
     #BLEND:
       // ========================================================================================================
       // Blending 
       // ========================================================================================================
       // Definition of blending (PathData: cmdParameters.bufferMode)
       // The parameter name is defined as "BLEND"
       // 
       // If "BLEND" was found, set the defined values in the connected PathData
       // The values are defined as "DirectValues" because the value to set is directly written here in this FC
       // Buffer mode (cmdParameters.bufferMode)
       // #parameterDefinition.directValues.cmdParameters.bufferMode := 5;
       // --> Set the bufferMode to 5 (Blending with high velocity)
       // 
       // Also set the priority #parameterDefinition.priorities.cmdParameters.bufferMode := "LKINLANG_PRIO_DEFINED";
       // 
       // Properties:
       // ----------
       // "LKINLANG_PRG_MODAL": Modal in program to save velocity value once set
       // 
       // Conditions:
       // ----------
       // Conditions are used to make other parameters mandatory.
       // Here the parameter "RADIUS" must be programmed the same line, because blending consits of the bufferMode and the TransitionParameter[1].
       // There can be up to "LKINLANG_NUMBER_OF_CONDITIONS" conditions.
       // How to configure:
       // 1. Set conditions[#tempConditionCounter].ParameterNumber to the parameter you want to check
       // 2. Set conditions[#tempConditionCounter].Mode according to where the parameter has to be written
       //    These modes are possible:
       //    "LKINLANG_CONDITION_IN_LINE" --> Selected parameter must be written in the same line
       //    "LKINLANG_CONDITION_IN_COMMAND" --> Selected parameter must be written in the same motion command
       //    "LKINLANG_CONDITION_IN_PROGRAM" --> Selected parameter must be written somewhere in the program before
       // 3. The setting #parameterDefinition.conditions[#tempConditionCounter].Group can be used to group parameters
       //    Only one condition of each group must be fulfilled.
       //    Also make sure groups are not used twice for other parameters; they must be unique
       //    
       // 
       // Parameter name definition
       #parameterDefinition.parameterNameString := 'BLEND';
       #parameterDefinition.parameterNameNumber := -1;

       // Matching to PathData
       #parameterDefinition.directValues.cmdParameters.bufferMode := 5; // BlendHigh

       // Priorities
       #parameterDefinition.priorities.cmdParameters.bufferMode := "LKINLANG_PRIO_DEFINED";

       // Properties
       #parameterDefinition.properties := "LKINLANG_PRG_MODAL";

       // Conditions
       #tempConditionCounter := 1;
       #parameterDefinition.conditions[#tempConditionCounter].ParameterNumber := #RADIUS;
       #parameterDefinition.conditions[#tempConditionCounter].Mode := "LKINLANG_CONDITION_IN_LINE";
       #parameterDefinition.conditions[#tempConditionCounter].Group := 10;

       // Valid counts per line
       #parameterDefinition.validCountPerLine := 1;
       // ========================================================================================================


     #RADIUS:
       // ========================================================================================================
       // Transition parameter
       // ========================================================================================================
       // Definition of TransitionParameter[1] (PathData: cmdParameters.transitionParameters[1])
       // The parameter name is defined as "R"
       // 
       // If "R" was found, set the defined values in the connected PathData
       // The value is defined as "FollowingValue" because the value is not written here, but in the program line after this parameter
       // e.g. R15 <-- 15 is taken as transitionParameter[1]
       // To do this, set #parameterDefinition.followingValues[1].cmdParameters.transitionParameters[1] := TRUE;
       // 
       // Also set the priority #parameterDefinition.priorities.cmdParameters.transitionParameters[1] := "LKINLANG_PRIO_DEFINED";
       // 
       // Properties:
       // ----------
       // "LKINLANG_PRG_MODAL": Modal in program to save transition parameter
       // 
       // Conditions:
       // ----------
       // This parameter is a condition for "BLEND", whenever "BLEND" is programmed, also "R" must be written in the same line.
       // See definition above.
       // 
       //
       // Parameter name definition
       #parameterDefinition.parameterNameString := 'R';
       #parameterDefinition.parameterNameNumber := -1;

       // Matching to PathData
       #parameterDefinition.followingValues[1].cmdParameters.transitionParameters[1] := TRUE; // Transition parameter [1] is set

       // Priorities
       #parameterDefinition.priorities.cmdParameters.transitionParameters[1] := "LKINLANG_PRIO_DEFINED";

       // Properties
       #parameterDefinition.properties := "LKINLANG_PRG_MODAL";

       // Valid counts per line
       #parameterDefinition.validCountPerLine := 1;
       // ========================================================================================================

       // ========================================================================================================
       // General Parameters
       // ========================================================================================================
     #X:
       // ========================================================================================================
       #parameterDefinition.parameterNameString := 'X';
       #parameterDefinition.parameterNameNumber := -1;
       #parameterDefinition.properties := "LKINLANG_CHECK_LIMITS" + "LKINLANG_EQUATION";
       #parameterDefinition.priorities.cmdCoordinates.cartesianPosition.x := "LKINLANG_PRIO_DEFINED";
       #parameterDefinition.followingValues[1].cmdCoordinates.cartesianPosition.x := true;
       // ========================================================================================================

     #Y:
       // ========================================================================================================
       #parameterDefinition.parameterNameString := 'Y';
       #parameterDefinition.parameterNameNumber := -1;
       #parameterDefinition.properties := "LKINLANG_CHECK_LIMITS" + "LKINLANG_EQUATION";
       #parameterDefinition.priorities.cmdCoordinates.cartesianPosition.y := "LKINLANG_PRIO_DEFINED";
       #parameterDefinition.followingValues[1].cmdCoordinates.cartesianPosition.y := true;
       // ========================================================================================================

     #Z:
       // ========================================================================================================
       #parameterDefinition.parameterNameString := 'Z';
       #parameterDefinition.parameterNameNumber := -1;
       #parameterDefinition.properties := "LKINLANG_CHECK_LIMITS" + "LKINLANG_EQUATION";
       #parameterDefinition.priorities.cmdCoordinates.cartesianPosition.z := "LKINLANG_PRIO_DEFINED";
       #parameterDefinition.followingValues[1].cmdCoordinates.cartesianPosition.z := true;
       // ========================================================================================================

     #END:
       // ========================================================================================================
       // End of program 
       // ========================================================================================================
       // This command is needed to signalize the end of a program
       // It is always necessary else the application will stay busy even without further program lines
       // ========================================================================================================
       // Parameter name definition
       #parameterDefinition.parameterNameString := 'END';
       #parameterDefinition.parameterNameNumber := -1;

       // Matching to PathData
       #parameterDefinition.directValues.cmdType := -1;

       // Priorities
       #parameterDefinition.priorities.cmdType := "LKINLANG_PRIO_DEFINED";

       // Properties
       #parameterDefinition.properties := "LKINLANG_MOTION_CMD";

       // Valid counts per line
       #parameterDefinition.validCountPerLine := 1;
       // ========================================================================================================

       // ========================================================================================================
       // Expand this list with more parameter definitions
       // ========================================================================================================
       // ...
       // ========================================================================================================
     ELSE
       // invalid case number
       #parameterNo := -2;

   END_CASE;
END_FUNCTION

// folder: LKinLang_Blocks/LKinLang_SubBlocks

FUNCTION "LKinLang_CalcMathAndBool" : "LKinLang_typeMathParserResult"   // FC35452, SCL
TITLE = LKinLang_CalcMathAndBool
{ S7_Optimized_Access := 'TRUE' }
AUTHOR : tech.team.motioncontrol@siemens.com
FAMILY : LKinLang
VERSION : 1.1
// This FC calculates math and boolean expressions / The FC to calculates math and boolean expressions
   VAR_INPUT
      inputString : String[254];   // Input string
   END_VAR
   VAR_TEMP
      tempCounter : Int;   // Temporary counter for length of the input string
      tempLenCodeline : Int;   // Temporary variable for length of the input string
      tempInputString : String[254];   // Temporary variable for input string
      tempLengthOfString : Int;   // Number of used signs in string
      tempPositionOfConvertedString : Int;   // Counter: Positon of converted character
      tempPositionOfPrePostfix : Int;   // Counter: Array PrePostfix
      tempPositionOfPostfix : Int;   // Counter: Postfix notation
      tempPositionOfOperatorStack : Int;   // Counter: Operator storage
      tempNumberOfMultiDigitNo : Int;   // Number of multi digits
      tempNumberOfBrackets : Int;   // Number of brackets
      tempDecimalPoint : Int;   // Monitoring only one comma per number
      tempDenominatorDecimalNumbers : LReal;   // Denominator for generating decimal number
      tempNumberOfNegBrackets : Int;   // Number of negative brackets
      tempNumberOfNegFunctions : Int;   // Number of negativ functions
      tempNumberOfDecimalNo : Int;   // Number of decimal numbers
      tempNumberOfNegTerm : Int;   // Number of negative expressions (brackets / functions)
      tempMaxPositionOfPrePostfix : Int;   // Max number of aPrePostfix array
      tempMaxOfPostfixPosition : Int;   // Max number of aPostfixNotation
      tempPositionOfIntermediateResult : Int;   // Counter: Interim results
      tempNextPostfixNumberIsNegative : Bool;   // Negative number detected
      tempStringConvertedToLReal : Array[0..#LGCODE_MTH_PRSR_STRING_LENGTH] of LReal;   // Converted numbers to LReal
      tempPrePostfix : Array[0..#LGCODE_MTH_PRSR_STRING_LENGTH] of LReal;   // Sign- and syntax check
      tempPostfixNotation : Array[0..#LGCODE_MTH_PRSR_STRING_LENGTH] of LReal;   // Postfix notation
      tempStackForOperators : Array[0..#LGCODE_MTH_PRSR_STRING_LENGTH] of LReal;   // Stack for operators
      tempPositionMultiDigitNumbers : Array[0..#LGCODE_MTH_PRSR_STRING_LENGTH] of Int;   // Positions of multi digits
      tempPositionOfNegBrackets : Array[0..#LGCODE_MTH_PRSR_STRING_LENGTH] of Int;   // Positions of opening brackets
      tempPositionOfNegFunctions : Array[0..#LGCODE_MTH_PRSR_STRING_LENGTH] of Int;   // Positions of negative math expressions
      tempPositionOfNegTerm : Array[0..#LGCODE_MTH_PRSR_STRING_LENGTH] of Int;   // Positions of negative expressions
      tempStackOfIntermediateResults : Array[0..#LGCODE_MTH_PRSR_STRING_LENGTH] of LReal;   // Stack for interim results
      tempPositionDecimalNumbers : Array[0..#LGCODE_MTH_PRSR_STRING_LENGTH] of Int;   // Position decimal numbers: Exponential calculation
   END_VAR
   // Ret_Val : Return values of function
   VAR CONSTANT
      LGCODE_MTH_PRSR_STRING_LENGTH : Int := 82;   // Maxumum string length of internal variables / Maxumum string length of internal varaibles
      LGCODE_MTH_PRSR_NO_ERR : DInt := 0;   // Error ID: No error
      LGCODE_MTH_PRSR_ERR_ID_INVALID_SYNTAX : DInt := 1;   // Error ID: Invalid syntax in string
      LGCODE_MTH_PRSR_ERR_ID_INVALID_CHARACTER : DInt := 2;   // Error ID: Invalid character in string
      LGCODE_MTH_PRSR_ERR_ID_NEAGTIVE_SQUARE_ROOT_ARGUMENT : DInt := 3;   // Error ID: Negative square root
      LGCODE_MTH_PRSR_ERR_ID_DIVISION_BY_ZERO : DInt := 4;   // Error ID: Division by zero
      LGCODE_MTH_PRSR_ERR_ID_BASIS_ZERO_EXPONENT_NEGATIVE : DInt := 5;   // Error ID: Basis is zero and exponent is negative
      LGCODE_MTH_PRSR_ERR_ID_BASIS_NEGATIVE_EXPONENT_REAL : DInt := 6;   // Error ID: Basis is negative and exponent is decimal
      LGCODE_MTH_PRSR_PI : LReal := 3.14159265358979;   // Mathconstant for Pi
      LGCODE_MTH_PRSR_NUMBER_0 : LReal := 48.0;   // Decimal value of '0'
      LGCODE_MTH_PRSR_NUMBER_1 : LReal := 49.0;   // Decimal value of '1'
      LGCODE_MTH_PRSR_NUMBER_2 : LReal := 50.0;   // Decimal value of '2'
      LGCODE_MTH_PRSR_NUMBER_3 : LReal := 51.0;   // Decimal value of '3'
      LGCODE_MTH_PRSR_NUMBER_4 : LReal := 52.0;   // Decimal value of '4'
      LGCODE_MTH_PRSR_NUMBER_5 : LReal := 53.0;   // Decimal value of '5'
      LGCODE_MTH_PRSR_NUMBER_6 : LReal := 54.0;   // Decimal value of '6'
      LGCODE_MTH_PRSR_NUMBER_7 : LReal := 55.0;   // Decimal value of '7'
      LGCODE_MTH_PRSR_NUMBER_8 : LReal := 56.0;   // Decimal value of '8'
      LGCODE_MTH_PRSR_NUMBER_9 : LReal := 57.0;   // Decimal value of '9'
      LGCODE_MTH_PRSR_UPPER_CASE_C : LReal := 67.0;   // Decimal value of 'C'
      LGCODE_MTH_PRSR_UPPER_CASE_I : LReal := 73.0;   // Decimal value of 'I'
      LGCODE_MTH_PRSR_UPPER_CASE_N : LReal := 78.0;   // Decimal value of 'N'
      LGCODE_MTH_PRSR_UPPER_CASE_O : LReal := 79.0;   // Decimal value of 'O'
      LGCODE_MTH_PRSR_UPPER_CASE_Q : LReal := 81.0;   // Decimal value of 'Q'
      LGCODE_MTH_PRSR_UPPER_CASE_R : LReal := 82.0;   // Decimal value of 'R'
      LGCODE_MTH_PRSR_UPPER_CASE_S : LReal := 83.0;   // Decimal value of 'S'
      LGCODE_MTH_PRSR_UPPER_CASE_T : LReal := 84.0;   // Decimal value of 'T'
      LGCODE_MTH_PRSR_LOWER_CASE_C : LReal := 99.0;   // Decimal value of 'c'
      LGCODE_MTH_PRSR_LOWER_CASE_I : LReal := 105.0;   // Decimal value of 'i'
      LGCODE_MTH_PRSR_LOWER_CASE_N : LReal := 110.0;   // Decimal value of 'n'
      LGCODE_MTH_PRSR_LOWER_CASE_O : LReal := 111.0;   // Decimal value of 'o'
      LGCODE_MTH_PRSR_LOWER_CASE_Q : LReal := 113.0;   // Decimal value of 'q'
      LGCODE_MTH_PRSR_LOWER_CASE_R : LReal := 114.0;   // Decimal value of 'r'
      LGCODE_MTH_PRSR_LOWER_CASE_S : LReal := 115.0;   // Decimal value of 's'
      LGCODE_MTH_PRSR_LOWER_CASE_T : LReal := 116.0;   // Decimal value of 't'
      LGCODE_MTH_PRSR_MULTIPLIER_FOR_MULTI_DIGIT_NO : LReal := 10.0;   // Decimal base
      LGCODE_MTH_PRSR_COSINUS : LReal := 34.0;   // internal constant for 'cos'
      LGCODE_MTH_PRSR_SQUARE : LReal := 35.0;   // internal constant for 'sqr'
      LGCODE_MTH_PRSR_SQUAREROOT : LReal := 36.0;   // internal constant for 'sqrt'
      LGCODE_MTH_PRSR_SINUS : LReal := 37.0;   // internal constant for 'sin'
      LGCODE_MTH_PRSR_OPEN_BRACKET : LReal := 40.0;   // Decimal value of '('
      LGCODE_MTH_PRSR_CLOSE_BRACKET : LReal := 41.0;   // Decimal value of ')'
      LGCODE_MTH_PRSR_TIMES : LReal := 42.0;   // Decimal value of '*'
      LGCODE_MTH_PRSR_PLUS : LReal := 43.0;   // Decimal value of '+'
      LGCODE_MTH_PRSR_MINUS : LReal := 45.0;   // Decimal value of '-'
      LGCODE_MTH_PRSR_DECIMAL_POINT : LReal := 46.0;   // Decimal value of '.'
      LGCODE_MTH_PRSR_DIVIDE : LReal := 47.0;   // Decimal value of '/'
      LGCODE_MTH_PRSR_TO_THE_POWER_OF : LReal := 94.0;   // Decimal value of '^'
      LGCODE_MTH_PRSR_CHAR_C : LReal := 99.0;   // Decimal value of 'c'
      LGCODE_MTH_PRSR_CHAR_I : LReal := 105.0;   // Decimal value of 'i'
      LGCODE_MTH_PRSR_CHAR_N : LReal := 110.0;   // Decimal value of 'n'
      LGCODE_MTH_PRSR_CHAR_O : LReal := 111.0;   // Decimal value of 'o'
      LGCODE_MTH_PRSR_CHAR_Q : LReal := 113.0;   // Decimal value of 'q'
      LGCODE_MTH_PRSR_CHAR_R : LReal := 114.0;   // Decimal value of 'r'
      LGCODE_MTH_PRSR_CHAR_S : LReal := 115.0;   // Decimal value of 's'
      LGCODE_MTH_PRSR_CHAR_T : LReal := 116.0;   // Decimal value of 't'
      LGCODE_MTH_PRSR_LOGICAL_NOT : LReal := 33.0;   // Decimal value of '!'
      LGCODE_MTH_PRSR_LOGICAL_AND : LReal := 38.0;   // Decimal value of '&'
      LGCODE_MTH_PRSR_LOGICAL_LESS : LReal := 60.0;   // Decimal value of '<'
      LGCODE_MTH_PRSR_LOGICAL_EQUAL : LReal := 61.0;   // Decimal value of '='
      LGCODE_MTH_PRSR_LOGICAL_GREATER : LReal := 62.0;   // Decimal value of '>'
      LGCODE_MTH_PRSR_LOGICAL_GREATER_EQUAL : LReal := 103.0;   // Decimal value of '>='
      LGCODE_MTH_PRSR_LOGICAL_LESS_EQUAL : LReal := 108.0;   // Decimal value of '<='
      LGCODE_MTH_PRSR_LOGICAL_OR : LReal := 124.0;   // Decimal value of '|'
      LGCODE_MTH_PRSR_LOGICAL_NOT_EQUAL : LReal := 156.0;   // Decimal value of '<>'
   END_VAR
BEGIN
   //==========================================================================================
   // SIEMENS AG
   // (c)Copyright 2019 All Rights Reserved
   //------------------------------------------------------------------------------------------
   // Library: LKinLang
   // Tested with: S7-1517T-3 PN/DP
   // Engineering: TIA Portal V15
   // Restrictions: ---
   // Requirements: S7-1500T FW 2.5
   // Functionality: LKinLang_CalcMathAndBool
   // The FC to calculates math and boolean expressions
   // 
   // Support: tech.team.motioncontrol@siemens.com
   // Note: Parameter comments are only available in language 'English (United States)'
   //------------------------------------------------------------------------------------------
   // Change log table:
   // Version    Date          Expert in charge    Changes applied
   // 02.02.00   28.05.2019    FR                  First version for SIMATIC  
   //===========================================================================================

   // Initialize temp variables
   #LKinLang_CalcMathAndBool.finalResult := 0;
   #tempLengthOfString:= 1;                      
   #tempPositionOfConvertedString := 1;                
   #tempPositionOfPrePostfix := 1;                 
   #tempPositionOfPrePostfix := 1;                 
   #tempPositionOfPostfix := 1;                 
   #tempPositionOfOperatorStack := 1;                 
   #tempNumberOfMultiDigitNo := 1;                 
   #tempNumberOfBrackets := 1;                 
   #tempDecimalPoint := 1;                 
   #tempDenominatorDecimalNumbers := 10.0;             
   #tempNumberOfNegBrackets := 1; 
   #tempNumberOfNegFunctions := 1;
   #tempNumberOfDecimalNo := 1;
   #tempNumberOfNegTerm := 1;
   #tempMaxPositionOfPrePostfix :=0;
   #tempMaxOfPostfixPosition :=0;
   #tempPositionOfIntermediateResult := 2;
   #tempNextPostfixNumberIsNegative := FALSE;

   // Get local copy of math string
   #tempInputString := #inputString;

   //======================================================================
   // Replace e in referenced ascii line with *10^
   // Sometimes you get something like this "2.33455e-10" by converting 
   // LREAL to STRING
   //======================================================================
   // Replace e by *10^ (It´s possible to get the e when you convert LREAL to String)
   #tempLenCodeline := LEN(#tempInputString);
   // Search e
   FOR #tempCounter := 1 TO #tempLenCodeline DO
     IF #tempInputString[#tempCounter] = '$65' THEN // e 
       // Replace e with *10^ (4digits)
       IF #tempLenCodeline <= 254 - 4 THEN
         #tempInputString := DELETE(IN := #tempInputString, L := 1, P := #tempCounter);
         #tempInputString := INSERT(IN1 := #tempInputString, IN2 := '*10^', P := #tempCounter - 1);
         #tempLenCodeline := LEN(#tempInputString);
       ELSE
         ;// not enough place in string
         #tempInputString := DELETE(IN := #tempInputString, L := 4, P := #tempCounter - 3);
         #tempInputString := INSERT(IN1 := #tempInputString, IN2 := '*10^', P := #tempCounter - 4);
         #tempLenCodeline := LEN(#tempInputString);
       END_IF;

     ELSE
       ; // No tap
     END_IF;
   END_FOR;
   // ------------------------------------------------------------------------------------------

   #tempLengthOfString := LEN(IN := #tempInputString);    // Get new length of string

   //Zeichenkontrolle
   //Codierungen in Zahlen umwandeln
   WHILE #tempPositionOfConvertedString <= #tempLengthOfString DO
     //String einlesen und nach LREAL konvertieren
     #tempStringConvertedToLReal[#tempPositionOfConvertedString] :=
     DINT_TO_LREAL(CHAR_TO_DINT(#tempInputString[#tempPositionOfConvertedString]));

     //Zeichenkontrolle
     IF    //Codierungen in Zahlen umwandeln
       #tempStringConvertedToLReal[#tempPositionOfConvertedString] = #LGCODE_MTH_PRSR_NUMBER_0
     THEN
       #tempPrePostfix[#tempPositionOfPrePostfix] := #LGCODE_MTH_PRSR_NUMBER_0;
       #tempPositionOfPrePostfix := #tempPositionOfPrePostfix + 1;
     ELSIF
       #tempStringConvertedToLReal[#tempPositionOfConvertedString] = #LGCODE_MTH_PRSR_NUMBER_1
     THEN
       #tempPrePostfix[#tempPositionOfPrePostfix] := #LGCODE_MTH_PRSR_NUMBER_1;
       #tempPositionOfPrePostfix := #tempPositionOfPrePostfix + 1;
     ELSIF
       #tempStringConvertedToLReal[#tempPositionOfConvertedString] = #LGCODE_MTH_PRSR_NUMBER_2
     THEN
       #tempPrePostfix[#tempPositionOfPrePostfix] := #LGCODE_MTH_PRSR_NUMBER_2;
       #tempPositionOfPrePostfix := #tempPositionOfPrePostfix + 1;
     ELSIF
       #tempStringConvertedToLReal[#tempPositionOfConvertedString] = #LGCODE_MTH_PRSR_NUMBER_3
     THEN
       #tempPrePostfix[#tempPositionOfPrePostfix] := #LGCODE_MTH_PRSR_NUMBER_3;
       #tempPositionOfPrePostfix := #tempPositionOfPrePostfix + 1;
     ELSIF
       #tempStringConvertedToLReal[#tempPositionOfConvertedString] = #LGCODE_MTH_PRSR_NUMBER_4
     THEN
       #tempPrePostfix[#tempPositionOfPrePostfix] := #LGCODE_MTH_PRSR_NUMBER_4;
       #tempPositionOfPrePostfix := #tempPositionOfPrePostfix + 1;
     ELSIF
       #tempStringConvertedToLReal[#tempPositionOfConvertedString] = #LGCODE_MTH_PRSR_NUMBER_5
     THEN
       #tempPrePostfix[#tempPositionOfPrePostfix] := #LGCODE_MTH_PRSR_NUMBER_5;
       #tempPositionOfPrePostfix := #tempPositionOfPrePostfix + 1;
     ELSIF
       #tempStringConvertedToLReal[#tempPositionOfConvertedString] = #LGCODE_MTH_PRSR_NUMBER_6
     THEN
       #tempPrePostfix[#tempPositionOfPrePostfix] := #LGCODE_MTH_PRSR_NUMBER_6;
       #tempPositionOfPrePostfix := #tempPositionOfPrePostfix + 1;
     ELSIF
       #tempStringConvertedToLReal[#tempPositionOfConvertedString] = #LGCODE_MTH_PRSR_NUMBER_7
     THEN
       #tempPrePostfix[#tempPositionOfPrePostfix] := #LGCODE_MTH_PRSR_NUMBER_7;
       #tempPositionOfPrePostfix := #tempPositionOfPrePostfix + 1;
     ELSIF
       #tempStringConvertedToLReal[#tempPositionOfConvertedString] = #LGCODE_MTH_PRSR_NUMBER_8
     THEN
       #tempPrePostfix[#tempPositionOfPrePostfix] := #LGCODE_MTH_PRSR_NUMBER_8;
       #tempPositionOfPrePostfix := #tempPositionOfPrePostfix + 1;
     ELSIF
       #tempStringConvertedToLReal[#tempPositionOfConvertedString] = #LGCODE_MTH_PRSR_NUMBER_9
     THEN
       #tempPrePostfix[#tempPositionOfPrePostfix] := #LGCODE_MTH_PRSR_NUMBER_9;
       #tempPositionOfPrePostfix := #tempPositionOfPrePostfix + 1;
     ELSIF
       //Größer-Gleich erzeugen
       (#tempStringConvertedToLReal[#tempPositionOfConvertedString - 1] = #LGCODE_MTH_PRSR_LOGICAL_GREATER) AND
       (#tempStringConvertedToLReal[#tempPositionOfConvertedString] = #LGCODE_MTH_PRSR_LOGICAL_EQUAL)
     THEN
       #tempPrePostfix[#tempPositionOfPrePostfix - 1] := #LGCODE_MTH_PRSR_LOGICAL_GREATER_EQUAL;
     ELSIF
       //Kleiner-Gleich erzeugen
       (#tempStringConvertedToLReal[#tempPositionOfConvertedString - 1] = #LGCODE_MTH_PRSR_LOGICAL_LESS) AND
       (#tempStringConvertedToLReal[#tempPositionOfConvertedString] = #LGCODE_MTH_PRSR_LOGICAL_EQUAL)
     THEN
       #tempPrePostfix[#tempPositionOfPrePostfix - 1] := #LGCODE_MTH_PRSR_LOGICAL_LESS_EQUAL;
     ELSIF
       //Ungleich erzeugen
       (#tempStringConvertedToLReal[#tempPositionOfConvertedString - 1] = #LGCODE_MTH_PRSR_LOGICAL_LESS) AND
       (#tempStringConvertedToLReal[#tempPositionOfConvertedString] = #LGCODE_MTH_PRSR_LOGICAL_GREATER)
     THEN
       #tempPrePostfix[#tempPositionOfPrePostfix - 1] := #LGCODE_MTH_PRSR_LOGICAL_NOT_EQUAL;
     ELSIF
       ((#tempStringConvertedToLReal[#tempPositionOfConvertedString] = #LGCODE_MTH_PRSR_UPPER_CASE_S) OR
       (#tempStringConvertedToLReal[#tempPositionOfConvertedString] = #LGCODE_MTH_PRSR_LOWER_CASE_S))
     THEN
       #tempPrePostfix[#tempPositionOfPrePostfix] := #LGCODE_MTH_PRSR_CHAR_S;
       #tempPositionOfPrePostfix := #tempPositionOfPrePostfix + 1;
     ELSIF
       ((#tempStringConvertedToLReal[#tempPositionOfConvertedString] = #LGCODE_MTH_PRSR_UPPER_CASE_I) OR
       (#tempStringConvertedToLReal[#tempPositionOfConvertedString] = #LGCODE_MTH_PRSR_LOWER_CASE_I))
     THEN
       #tempPrePostfix[#tempPositionOfPrePostfix] := #LGCODE_MTH_PRSR_CHAR_I;
       #tempPositionOfPrePostfix := #tempPositionOfPrePostfix + 1;
     ELSIF
       ((#tempStringConvertedToLReal[#tempPositionOfConvertedString] = #LGCODE_MTH_PRSR_UPPER_CASE_N) OR
       (#tempStringConvertedToLReal[#tempPositionOfConvertedString] = #LGCODE_MTH_PRSR_LOWER_CASE_N))
     THEN
       #tempPrePostfix[#tempPositionOfPrePostfix] := #LGCODE_MTH_PRSR_CHAR_N;
       #tempPositionOfPrePostfix := #tempPositionOfPrePostfix + 1;
     ELSIF
       ((#tempStringConvertedToLReal[#tempPositionOfConvertedString] = #LGCODE_MTH_PRSR_UPPER_CASE_C) OR
       (#tempStringConvertedToLReal[#tempPositionOfConvertedString] = #LGCODE_MTH_PRSR_LOWER_CASE_C))
     THEN
       #tempPrePostfix[#tempPositionOfPrePostfix] := #LGCODE_MTH_PRSR_CHAR_C;
       #tempPositionOfPrePostfix := #tempPositionOfPrePostfix + 1;
     ELSIF
       ((#tempStringConvertedToLReal[#tempPositionOfConvertedString] = #LGCODE_MTH_PRSR_UPPER_CASE_O) OR
       (#tempStringConvertedToLReal[#tempPositionOfConvertedString] = #LGCODE_MTH_PRSR_LOWER_CASE_O))
     THEN
       #tempPrePostfix[#tempPositionOfPrePostfix] := #LGCODE_MTH_PRSR_CHAR_O;
       #tempPositionOfPrePostfix := #tempPositionOfPrePostfix + 1;
     ELSIF
       ((#tempStringConvertedToLReal[#tempPositionOfConvertedString] = #LGCODE_MTH_PRSR_UPPER_CASE_Q) OR
       (#tempStringConvertedToLReal[#tempPositionOfConvertedString] = #LGCODE_MTH_PRSR_LOWER_CASE_Q))
     THEN
       #tempPrePostfix[#tempPositionOfPrePostfix] := #LGCODE_MTH_PRSR_CHAR_Q;
       #tempPositionOfPrePostfix := #tempPositionOfPrePostfix + 1;
     ELSIF
       ((#tempStringConvertedToLReal[#tempPositionOfConvertedString] = #LGCODE_MTH_PRSR_UPPER_CASE_R) OR
       (#tempStringConvertedToLReal[#tempPositionOfConvertedString] = #LGCODE_MTH_PRSR_LOWER_CASE_R))
     THEN
       #tempPrePostfix[#tempPositionOfPrePostfix] := #LGCODE_MTH_PRSR_CHAR_R;
       #tempPositionOfPrePostfix := #tempPositionOfPrePostfix + 1;
     ELSIF
       ((#tempStringConvertedToLReal[#tempPositionOfConvertedString] = #LGCODE_MTH_PRSR_UPPER_CASE_T) OR
       (#tempStringConvertedToLReal[#tempPositionOfConvertedString] = #LGCODE_MTH_PRSR_LOWER_CASE_T))
     THEN
       #tempPrePostfix[#tempPositionOfPrePostfix] := #LGCODE_MTH_PRSR_CHAR_T;
       #tempPositionOfPrePostfix := #tempPositionOfPrePostfix + 1;
     ELSIF
       ((#tempStringConvertedToLReal[#tempPositionOfConvertedString] = #LGCODE_MTH_PRSR_DECIMAL_POINT) OR
       (#tempStringConvertedToLReal[#tempPositionOfConvertedString] = #LGCODE_MTH_PRSR_OPEN_BRACKET) OR
       (#tempStringConvertedToLReal[#tempPositionOfConvertedString] = #LGCODE_MTH_PRSR_CLOSE_BRACKET) OR
       (#tempStringConvertedToLReal[#tempPositionOfConvertedString] = #LGCODE_MTH_PRSR_PLUS) OR
       (#tempStringConvertedToLReal[#tempPositionOfConvertedString] = #LGCODE_MTH_PRSR_MINUS) OR
       (#tempStringConvertedToLReal[#tempPositionOfConvertedString] = #LGCODE_MTH_PRSR_TIMES) OR
       (#tempStringConvertedToLReal[#tempPositionOfConvertedString] = #LGCODE_MTH_PRSR_DIVIDE) OR
       (#tempStringConvertedToLReal[#tempPositionOfConvertedString] = #LGCODE_MTH_PRSR_LOGICAL_GREATER) OR
       (#tempStringConvertedToLReal[#tempPositionOfConvertedString] = #LGCODE_MTH_PRSR_LOGICAL_LESS) OR
       (#tempStringConvertedToLReal[#tempPositionOfConvertedString] = #LGCODE_MTH_PRSR_LOGICAL_NOT) OR
       (#tempStringConvertedToLReal[#tempPositionOfConvertedString] = #LGCODE_MTH_PRSR_LOGICAL_EQUAL) OR
       (#tempStringConvertedToLReal[#tempPositionOfConvertedString] = #LGCODE_MTH_PRSR_LOGICAL_AND) OR
       (#tempStringConvertedToLReal[#tempPositionOfConvertedString] = #LGCODE_MTH_PRSR_LOGICAL_OR) OR
       (#tempStringConvertedToLReal[#tempPositionOfConvertedString] = #LGCODE_MTH_PRSR_OPEN_BRACKET) OR
       (#tempStringConvertedToLReal[#tempPositionOfConvertedString] = #LGCODE_MTH_PRSR_CLOSE_BRACKET) OR
       (#tempStringConvertedToLReal[#tempPositionOfConvertedString] = #LGCODE_MTH_PRSR_DECIMAL_POINT) OR
       (#tempStringConvertedToLReal[#tempPositionOfConvertedString] = #LGCODE_MTH_PRSR_LOGICAL_NOT) OR
       (#tempStringConvertedToLReal[#tempPositionOfConvertedString] = #LGCODE_MTH_PRSR_MINUS) OR
       (#tempStringConvertedToLReal[#tempPositionOfConvertedString] = #LGCODE_MTH_PRSR_TO_THE_POWER_OF))

     THEN
       #tempPrePostfix[#tempPositionOfPrePostfix] := #tempStringConvertedToLReal[#tempPositionOfConvertedString];
       #tempPositionOfPrePostfix := #tempPositionOfPrePostfix + 1;
     ELSE    //Unzulässiges Zeichen
       #LKinLang_CalcMathAndBool.errorID := #LGCODE_MTH_PRSR_ERR_ID_INVALID_CHARACTER;
       #LKinLang_CalcMathAndBool.finalResult:= 0;

       RETURN;
     END_IF;
     #tempPositionOfConvertedString := #tempPositionOfConvertedString + 1;
     #tempMaxPositionOfPrePostfix := #tempPositionOfPrePostfix - 1;
   END_WHILE;

   //Syntaxkontrolle
   #tempPositionOfPrePostfix := 1;
   WHILE #tempPositionOfPrePostfix <= #tempMaxPositionOfPrePostfix DO
     //Zahl und nächstes Zeichen Zahl/schließende Klammer/Dezimalpunkt/boolescher Operator/
     //mathematischer Operator oder Ende STRING dann OK
     IF ((#tempPrePostfix[#tempPositionOfPrePostfix] >= #LGCODE_MTH_PRSR_NUMBER_0) AND
       (#tempPrePostfix[#tempPositionOfPrePostfix] <= #LGCODE_MTH_PRSR_NUMBER_9)) AND
       (((#tempPrePostfix[#tempPositionOfPrePostfix + 1] >= #LGCODE_MTH_PRSR_NUMBER_0) AND
       (#tempPrePostfix[#tempPositionOfPrePostfix + 1] <= #LGCODE_MTH_PRSR_NUMBER_9)) OR
       (#tempPrePostfix[#tempPositionOfPrePostfix + 1] = #LGCODE_MTH_PRSR_DECIMAL_POINT) OR
       (#tempPrePostfix[#tempPositionOfPrePostfix + 1] = #LGCODE_MTH_PRSR_CLOSE_BRACKET) OR
       (#tempPrePostfix[#tempPositionOfPrePostfix + 1] = #LGCODE_MTH_PRSR_PLUS) OR
       (#tempPrePostfix[#tempPositionOfPrePostfix + 1] = #LGCODE_MTH_PRSR_MINUS) OR
       (#tempPrePostfix[#tempPositionOfPrePostfix + 1] = #LGCODE_MTH_PRSR_TIMES) OR
       (#tempPrePostfix[#tempPositionOfPrePostfix + 1] = #LGCODE_MTH_PRSR_DIVIDE) OR
       (#tempPrePostfix[#tempPositionOfPrePostfix + 1] = #LGCODE_MTH_PRSR_DECIMAL_POINT) OR
       (#tempPrePostfix[#tempPositionOfPrePostfix + 1] = #LGCODE_MTH_PRSR_CLOSE_BRACKET) OR
       (#tempPrePostfix[#tempPositionOfPrePostfix + 1] = #LGCODE_MTH_PRSR_LOGICAL_GREATER) OR
       (#tempPrePostfix[#tempPositionOfPrePostfix + 1] = #LGCODE_MTH_PRSR_LOGICAL_LESS) OR
       (#tempPrePostfix[#tempPositionOfPrePostfix + 1] = #LGCODE_MTH_PRSR_LOGICAL_EQUAL) OR
       (#tempPrePostfix[#tempPositionOfPrePostfix + 1] = #LGCODE_MTH_PRSR_LOGICAL_AND) OR
       (#tempPrePostfix[#tempPositionOfPrePostfix + 1] = #LGCODE_MTH_PRSR_LOGICAL_OR) OR
       (#tempPrePostfix[#tempPositionOfPrePostfix + 1] = #LGCODE_MTH_PRSR_LOGICAL_GREATER_EQUAL) OR
       (#tempPrePostfix[#tempPositionOfPrePostfix + 1] = #LGCODE_MTH_PRSR_LOGICAL_LESS_EQUAL) OR
       (#tempPrePostfix[#tempPositionOfPrePostfix + 1] = #LGCODE_MTH_PRSR_LOGICAL_NOT_EQUAL) OR
       (#tempPrePostfix[#tempPositionOfPrePostfix + 1] = #LGCODE_MTH_PRSR_TO_THE_POWER_OF) OR
       (#tempPositionOfPrePostfix = #tempMaxPositionOfPrePostfix))
     THEN
       ;
     ELSIF
       //MAL und nächstes Zeichen Zahl/Klammerauf/Minus/c/(s und dann (i oder q)) und nicht Ende dann OK
       (#tempPrePostfix[#tempPositionOfPrePostfix] = #LGCODE_MTH_PRSR_TIMES) AND
       (((#tempPrePostfix[#tempPositionOfPrePostfix + 1] >= #LGCODE_MTH_PRSR_NUMBER_0) AND
       (#tempPrePostfix[#tempPositionOfPrePostfix + 1] <= #LGCODE_MTH_PRSR_NUMBER_9)) OR
       (#tempPrePostfix[#tempPositionOfPrePostfix + 1] = #LGCODE_MTH_PRSR_LOGICAL_NOT) OR
       (#tempPrePostfix[#tempPositionOfPrePostfix + 1] = #LGCODE_MTH_PRSR_OPEN_BRACKET) OR
       (#tempPrePostfix[#tempPositionOfPrePostfix + 1] = #LGCODE_MTH_PRSR_MINUS) OR
       (#tempPrePostfix[#tempPositionOfPrePostfix + 1] = #LGCODE_MTH_PRSR_CHAR_C) OR
       ((#tempPrePostfix[#tempPositionOfPrePostfix + 1] = #LGCODE_MTH_PRSR_CHAR_S) AND
       ((#tempPrePostfix[#tempPositionOfPrePostfix + 2] = #LGCODE_MTH_PRSR_CHAR_I) OR
       (#tempPrePostfix[#tempPositionOfPrePostfix + 2] = #LGCODE_MTH_PRSR_CHAR_Q)))) AND
       (#tempPositionOfPrePostfix <> #tempMaxPositionOfPrePostfix)
     THEN
       IF #tempDecimalPoint > 1 THEN
         #tempDecimalPoint := #tempDecimalPoint - 1;
       END_IF;
     ELSIF
       //GETEILT und nächstes Zeichen Zahl/Klammerauf/Minus/c/(s und dann (i oder q)) und nicht Ende dann OK
       (#tempPrePostfix[#tempPositionOfPrePostfix] = #LGCODE_MTH_PRSR_DIVIDE) AND
       (((#tempPrePostfix[#tempPositionOfPrePostfix + 1] >= #LGCODE_MTH_PRSR_NUMBER_0) AND
       (#tempPrePostfix[#tempPositionOfPrePostfix + 1] <= #LGCODE_MTH_PRSR_NUMBER_9)) OR
       (#tempPrePostfix[#tempPositionOfPrePostfix + 1] = #LGCODE_MTH_PRSR_LOGICAL_NOT) OR
       (#tempPrePostfix[#tempPositionOfPrePostfix + 1] = #LGCODE_MTH_PRSR_OPEN_BRACKET) OR
       (#tempPrePostfix[#tempPositionOfPrePostfix + 1] = #LGCODE_MTH_PRSR_MINUS) OR
       (#tempPrePostfix[#tempPositionOfPrePostfix + 1] = #LGCODE_MTH_PRSR_CHAR_C) OR
       ((#tempPrePostfix[#tempPositionOfPrePostfix + 1] = #LGCODE_MTH_PRSR_CHAR_S) AND
       ((#tempPrePostfix[#tempPositionOfPrePostfix + 2] = #LGCODE_MTH_PRSR_CHAR_I) OR
       (#tempPrePostfix[#tempPositionOfPrePostfix + 2] = #LGCODE_MTH_PRSR_CHAR_Q)))) AND
       (#tempPositionOfPrePostfix <> #tempMaxPositionOfPrePostfix)
     THEN
       IF #tempDecimalPoint > 1 THEN
         #tempDecimalPoint := #tempDecimalPoint - 1;
       END_IF;
     ELSIF
       //PLUS und nächstes Zeichen Zahl/Klammerauf/Minus/c/(s und dann (i oder q)) und nicht Ende dann OK
       (#tempPrePostfix[#tempPositionOfPrePostfix] = #LGCODE_MTH_PRSR_PLUS) AND
       (((#tempPrePostfix[#tempPositionOfPrePostfix + 1] >= #LGCODE_MTH_PRSR_NUMBER_0) AND
       (#tempPrePostfix[#tempPositionOfPrePostfix + 1] <= #LGCODE_MTH_PRSR_NUMBER_9)) OR
       (#tempPrePostfix[#tempPositionOfPrePostfix + 1] = #LGCODE_MTH_PRSR_LOGICAL_NOT) OR
       (#tempPrePostfix[#tempPositionOfPrePostfix + 1] = #LGCODE_MTH_PRSR_OPEN_BRACKET) OR
       (#tempPrePostfix[#tempPositionOfPrePostfix + 1] = #LGCODE_MTH_PRSR_MINUS) OR
       (#tempPrePostfix[#tempPositionOfPrePostfix + 1] = #LGCODE_MTH_PRSR_CHAR_C) OR
       ((#tempPrePostfix[#tempPositionOfPrePostfix + 1] = #LGCODE_MTH_PRSR_CHAR_S) AND
       ((#tempPrePostfix[#tempPositionOfPrePostfix + 2] = #LGCODE_MTH_PRSR_CHAR_I) OR
       (#tempPrePostfix[#tempPositionOfPrePostfix + 2] = #LGCODE_MTH_PRSR_CHAR_Q)))) AND
       (#tempPositionOfPrePostfix <> #tempMaxPositionOfPrePostfix)
     THEN
       IF #tempDecimalPoint > 1 THEN
         #tempDecimalPoint := #tempDecimalPoint - 1;
       END_IF;
     ELSIF
       //MINUS und nächstes Zeichen Zahl/Klammerauf/Minus/c/(s und dann (i oder q)) und nicht Ende dann OK
       (#tempPrePostfix[#tempPositionOfPrePostfix] = #LGCODE_MTH_PRSR_MINUS) AND
       (((#tempPrePostfix[#tempPositionOfPrePostfix + 1] >= #LGCODE_MTH_PRSR_NUMBER_0) AND
       (#tempPrePostfix[#tempPositionOfPrePostfix + 1] <= #LGCODE_MTH_PRSR_NUMBER_9)) OR
       (#tempPrePostfix[#tempPositionOfPrePostfix + 1] = #LGCODE_MTH_PRSR_LOGICAL_NOT) OR
       (#tempPrePostfix[#tempPositionOfPrePostfix + 1] = #LGCODE_MTH_PRSR_OPEN_BRACKET) OR

       ((#tempPrePostfix[#tempPositionOfPrePostfix + 1] = #LGCODE_MTH_PRSR_MINUS) AND
       (#tempPrePostfix[#tempPositionOfPrePostfix + 2] <> #LGCODE_MTH_PRSR_MINUS)) OR

       (#tempPrePostfix[#tempPositionOfPrePostfix + 1] = #LGCODE_MTH_PRSR_CHAR_C) OR
       ((#tempPrePostfix[#tempPositionOfPrePostfix + 1] = #LGCODE_MTH_PRSR_CHAR_S) AND
       ((#tempPrePostfix[#tempPositionOfPrePostfix + 2] = #LGCODE_MTH_PRSR_CHAR_I) OR
       (#tempPrePostfix[#tempPositionOfPrePostfix + 2] = #LGCODE_MTH_PRSR_CHAR_Q)))) AND
       (#tempPositionOfPrePostfix <> #tempMaxPositionOfPrePostfix)
     THEN
       IF #tempDecimalPoint > 1 THEN
         #tempDecimalPoint := #tempDecimalPoint - 1;
       END_IF;
     ELSIF
       //KOMMA und nächstes Zeichen Zahl dann OK
       (#tempPrePostfix[#tempPositionOfPrePostfix] = #LGCODE_MTH_PRSR_DECIMAL_POINT) AND
       (#tempPrePostfix[#tempPositionOfPrePostfix + 1] >= #LGCODE_MTH_PRSR_NUMBER_0) AND
       (#tempPrePostfix[#tempPositionOfPrePostfix + 1] <= #LGCODE_MTH_PRSR_NUMBER_9) AND
       (#tempPositionOfPrePostfix <> #tempMaxPositionOfPrePostfix) AND
       (#tempPositionOfPrePostfix > 1)
     THEN
       #tempDecimalPoint := #tempDecimalPoint + 1;
     ELSIF
       //s und nächstes Zeichen i oder q oder Klammerauf oder Minus oder Zahl und nicht Ende String dann OK
       (#tempPrePostfix[#tempPositionOfPrePostfix] = #LGCODE_MTH_PRSR_CHAR_S) AND
       ((#tempPrePostfix[#tempPositionOfPrePostfix + 1] = #LGCODE_MTH_PRSR_CHAR_I) OR
       (#tempPrePostfix[#tempPositionOfPrePostfix + 1] = #LGCODE_MTH_PRSR_CHAR_Q) OR
       (#tempPrePostfix[#tempPositionOfPrePostfix + 1] = #LGCODE_MTH_PRSR_OPEN_BRACKET) OR
       (#tempPrePostfix[#tempPositionOfPrePostfix + 1] = #LGCODE_MTH_PRSR_LOGICAL_NOT) OR
       (#tempPrePostfix[#tempPositionOfPrePostfix + 1] = #LGCODE_MTH_PRSR_MINUS) OR
       ((#tempPrePostfix[#tempPositionOfPrePostfix + 1] >= #LGCODE_MTH_PRSR_NUMBER_0) AND
       (#tempPrePostfix[#tempPositionOfPrePostfix + 1] <= #LGCODE_MTH_PRSR_NUMBER_9))) AND
       (#tempPositionOfPrePostfix <> #tempMaxPositionOfPrePostfix)
     THEN
       ;
     ELSIF
       //q und nächstes Zeichen r dann OK
       (#tempPrePostfix[#tempPositionOfPrePostfix] = #LGCODE_MTH_PRSR_CHAR_Q) AND (#tempPrePostfix[#tempPositionOfPrePostfix + 1] = #LGCODE_MTH_PRSR_CHAR_R)
     THEN
       ;
     ELSIF
       //r und nächstes Zeichen t oder oder Klammerauf oder Minus oder Zahl und nicht Ende String dann OK
       (#tempPrePostfix[#tempPositionOfPrePostfix] = #LGCODE_MTH_PRSR_CHAR_R) AND
       ((#tempPrePostfix[#tempPositionOfPrePostfix + 1] = #LGCODE_MTH_PRSR_CHAR_T) OR
       (#tempPrePostfix[#tempPositionOfPrePostfix + 1] = #LGCODE_MTH_PRSR_OPEN_BRACKET) OR
       (#tempPrePostfix[#tempPositionOfPrePostfix + 1] = #LGCODE_MTH_PRSR_MINUS) OR
       (#tempPrePostfix[#tempPositionOfPrePostfix + 1] = #LGCODE_MTH_PRSR_LOGICAL_NOT) OR
       ((#tempPrePostfix[#tempPositionOfPrePostfix + 1] >= #LGCODE_MTH_PRSR_NUMBER_0) AND
       (#tempPrePostfix[#tempPositionOfPrePostfix + 1] <= #LGCODE_MTH_PRSR_NUMBER_9))) AND
       (#tempPositionOfPrePostfix <> #tempMaxPositionOfPrePostfix)
     THEN
       ;
     ELSIF
       //t und nächstes Zeichen Zahl oder Klammerauf und nicht Ende String dann OK
       (#tempPrePostfix[#tempPositionOfPrePostfix] = #LGCODE_MTH_PRSR_CHAR_T) AND
       ((#tempPrePostfix[#tempPositionOfPrePostfix + 1] >= #LGCODE_MTH_PRSR_NUMBER_0) AND
       (#tempPrePostfix[#tempPositionOfPrePostfix + 1] <= #LGCODE_MTH_PRSR_NUMBER_9) OR
       (#tempPrePostfix[#tempPositionOfPrePostfix + 1] = #LGCODE_MTH_PRSR_OPEN_BRACKET) OR
       (#tempPrePostfix[#tempPositionOfPrePostfix + 1] = #LGCODE_MTH_PRSR_LOGICAL_NOT) OR
       (#tempPrePostfix[#tempPositionOfPrePostfix + 1] = #LGCODE_MTH_PRSR_MINUS)) AND
       (#tempPositionOfPrePostfix <> #tempMaxPositionOfPrePostfix)
     THEN
       ;
     ELSIF
       //c und nächstes Zeichen o dann OK
       (#tempPrePostfix[#tempPositionOfPrePostfix] = #LGCODE_MTH_PRSR_CHAR_C) AND (#tempPrePostfix[#tempPositionOfPrePostfix + 1] = #LGCODE_MTH_PRSR_CHAR_O)
     THEN
       ;
     ELSIF
       //o und nächstes Zeichen s dann OK
       (#tempPrePostfix[#tempPositionOfPrePostfix] = #LGCODE_MTH_PRSR_CHAR_O) AND (#tempPrePostfix[#tempPositionOfPrePostfix + 1] = #LGCODE_MTH_PRSR_CHAR_S)
     THEN
       ;
     ELSIF
       //i und nächstes Zeichen n dann OK
       (#tempPrePostfix[#tempPositionOfPrePostfix] = #LGCODE_MTH_PRSR_CHAR_I) AND (#tempPrePostfix[#tempPositionOfPrePostfix + 1] = #LGCODE_MTH_PRSR_CHAR_N)
     THEN
       ;
     ELSIF
       //n und nächstes Zeichen Zahl oder Klammerauf oder Minus und nicht Ende String dann OK
       (#tempPrePostfix[#tempPositionOfPrePostfix] = #LGCODE_MTH_PRSR_CHAR_N) AND
       (((#tempPrePostfix[#tempPositionOfPrePostfix + 1] >= #LGCODE_MTH_PRSR_NUMBER_0) AND
       (#tempPrePostfix[#tempPositionOfPrePostfix + 1] <= #LGCODE_MTH_PRSR_NUMBER_9)) OR
       (#tempPrePostfix[#tempPositionOfPrePostfix + 1] = #LGCODE_MTH_PRSR_OPEN_BRACKET) OR
       (#tempPrePostfix[#tempPositionOfPrePostfix + 1] = #LGCODE_MTH_PRSR_LOGICAL_NOT) OR
       (#tempPrePostfix[#tempPositionOfPrePostfix + 1] = #LGCODE_MTH_PRSR_MINUS)) AND
       (#tempPositionOfPrePostfix <> #tempMaxPositionOfPrePostfix)
     THEN
       ;
     ELSIF
       //Boolescher Operator und nächstes Zeichen Zahl/öffnende Klammerauf/Minus/NOT und nicht Ende dann OK
       ((#tempPrePostfix[#tempPositionOfPrePostfix] = #LGCODE_MTH_PRSR_LOGICAL_OR) OR
       (#tempPrePostfix[#tempPositionOfPrePostfix] = #LGCODE_MTH_PRSR_LOGICAL_AND) OR
       (#tempPrePostfix[#tempPositionOfPrePostfix] = #LGCODE_MTH_PRSR_LOGICAL_GREATER) OR
       (#tempPrePostfix[#tempPositionOfPrePostfix] = #LGCODE_MTH_PRSR_LOGICAL_LESS) OR
       (#tempPrePostfix[#tempPositionOfPrePostfix] = #LGCODE_MTH_PRSR_LOGICAL_EQUAL) OR
       (#tempPrePostfix[#tempPositionOfPrePostfix] = #LGCODE_MTH_PRSR_LOGICAL_GREATER_EQUAL) OR
       (#tempPrePostfix[#tempPositionOfPrePostfix] = #LGCODE_MTH_PRSR_LOGICAL_LESS_EQUAL) OR
       (#tempPrePostfix[#tempPositionOfPrePostfix] = #LGCODE_MTH_PRSR_LOGICAL_NOT_EQUAL))
       AND
       (((#tempPrePostfix[#tempPositionOfPrePostfix + 1] >= #LGCODE_MTH_PRSR_NUMBER_0) AND
       (#tempPrePostfix[#tempPositionOfPrePostfix + 1] <= #LGCODE_MTH_PRSR_NUMBER_9)) OR
       (#tempPrePostfix[#tempPositionOfPrePostfix + 1] = #LGCODE_MTH_PRSR_OPEN_BRACKET) OR
       (#tempPrePostfix[#tempPositionOfPrePostfix + 1] = #LGCODE_MTH_PRSR_LOGICAL_NOT) OR
       (#tempPrePostfix[#tempPositionOfPrePostfix + 1] = #LGCODE_MTH_PRSR_MINUS) OR
       (#tempPrePostfix[#tempPositionOfPrePostfix + 1] = #LGCODE_MTH_PRSR_CHAR_C) OR
       ((#tempPrePostfix[#tempPositionOfPrePostfix + 1] = #LGCODE_MTH_PRSR_CHAR_S) AND
       ((#tempPrePostfix[#tempPositionOfPrePostfix + 2] = #LGCODE_MTH_PRSR_CHAR_I) OR
       (#tempPrePostfix[#tempPositionOfPrePostfix + 2] = #LGCODE_MTH_PRSR_CHAR_Q))))
       AND
       (#tempPositionOfPrePostfix <> #tempMaxPositionOfPrePostfix)
     THEN
       IF #tempDecimalPoint > 1 THEN
         #tempDecimalPoint := #tempDecimalPoint - 1;
       END_IF;
     ELSIF
       //Exponetial-Operator und danach Zahl/Funktion/öffnende Klammer/
       //oder Minus (mit anschließender Funktion oder Zahl)
       ((#tempPrePostfix[#tempPositionOfPrePostfix] = #LGCODE_MTH_PRSR_TO_THE_POWER_OF)
       AND
       (((#tempPrePostfix[#tempPositionOfPrePostfix + 1] >= #LGCODE_MTH_PRSR_NUMBER_0) AND
       (#tempPrePostfix[#tempPositionOfPrePostfix + 1] <= #LGCODE_MTH_PRSR_NUMBER_9)) OR
       (#tempPrePostfix[#tempPositionOfPrePostfix + 1] = #LGCODE_MTH_PRSR_OPEN_BRACKET) OR
       (#tempPrePostfix[#tempPositionOfPrePostfix + 1] = #LGCODE_MTH_PRSR_MINUS) OR
       (#tempPrePostfix[#tempPositionOfPrePostfix + 1] = #LGCODE_MTH_PRSR_LOGICAL_NOT) OR
       (#tempPrePostfix[#tempPositionOfPrePostfix + 1] = #LGCODE_MTH_PRSR_CHAR_C) OR
       ((#tempPrePostfix[#tempPositionOfPrePostfix + 1] = #LGCODE_MTH_PRSR_CHAR_S) AND
       ((#tempPrePostfix[#tempPositionOfPrePostfix + 2] = #LGCODE_MTH_PRSR_CHAR_I) OR
       (#tempPrePostfix[#tempPositionOfPrePostfix + 2] = #LGCODE_MTH_PRSR_CHAR_Q)))
       AND
       (#tempPositionOfPrePostfix <> #tempMaxPositionOfPrePostfix)))
     THEN
       IF #tempDecimalPoint > 1 THEN
         #tempDecimalPoint := #tempDecimalPoint - 1;
       END_IF;
     ELSIF
       //NOT Operator und nächstes Zeichen eine Zahl oder eine öffnende Klammer und nicht Ende dann OK
       (#tempPrePostfix[#tempPositionOfPrePostfix] = #LGCODE_MTH_PRSR_LOGICAL_NOT)
       AND
       (((#tempPrePostfix[#tempPositionOfPrePostfix + 1] >= #LGCODE_MTH_PRSR_NUMBER_0) AND
       (#tempPrePostfix[#tempPositionOfPrePostfix + 1] <= #LGCODE_MTH_PRSR_NUMBER_9)) OR
       (#tempPrePostfix[#tempPositionOfPrePostfix + 1] = #LGCODE_MTH_PRSR_OPEN_BRACKET)
       AND
       (#tempPositionOfPrePostfix <> #tempMaxPositionOfPrePostfix))
     THEN
       ;
     ELSIF
       //Klammerauf und nächstes Zeichen Minus/Plus/öffnende Klammer/s/c oder Zahl dann OK
       (#tempPrePostfix[#tempPositionOfPrePostfix] = #LGCODE_MTH_PRSR_OPEN_BRACKET) AND
       ((#tempPrePostfix[#tempPositionOfPrePostfix + 1] = #LGCODE_MTH_PRSR_MINUS) OR
       (#tempPrePostfix[#tempPositionOfPrePostfix + 1] = #LGCODE_MTH_PRSR_OPEN_BRACKET) OR
       (#tempPrePostfix[#tempPositionOfPrePostfix + 1] = #LGCODE_MTH_PRSR_CHAR_S) OR
       (#tempPrePostfix[#tempPositionOfPrePostfix + 1] = #LGCODE_MTH_PRSR_CHAR_C) OR
       ((#tempPrePostfix[#tempPositionOfPrePostfix + 1] >= #LGCODE_MTH_PRSR_NUMBER_0) AND
       (#tempPrePostfix[#tempPositionOfPrePostfix + 1] <= #LGCODE_MTH_PRSR_NUMBER_9)))
     THEN
       #tempNumberOfBrackets := #tempNumberOfBrackets + 1;
     ELSIF
       //schließende Klammer und nächstes Zeichen schließende Klammer/pPlus/Minus/Mal/Geteilt/
       //boolescher Operator oder Ende STRING dann OK
       (#tempPrePostfix[#tempPositionOfPrePostfix] = #LGCODE_MTH_PRSR_CLOSE_BRACKET) AND
       ((#tempPrePostfix[#tempPositionOfPrePostfix + 1] = #LGCODE_MTH_PRSR_LOGICAL_OR) OR
       (#tempPrePostfix[#tempPositionOfPrePostfix + 1] = #LGCODE_MTH_PRSR_LOGICAL_AND) OR
       (#tempPrePostfix[#tempPositionOfPrePostfix + 1] = #LGCODE_MTH_PRSR_LOGICAL_GREATER) OR
       (#tempPrePostfix[#tempPositionOfPrePostfix + 1] = #LGCODE_MTH_PRSR_LOGICAL_LESS) OR
       (#tempPrePostfix[#tempPositionOfPrePostfix + 1] = #LGCODE_MTH_PRSR_LOGICAL_EQUAL) OR
       (#tempPrePostfix[#tempPositionOfPrePostfix + 1] = #LGCODE_MTH_PRSR_LOGICAL_NOT) OR
       (#tempPrePostfix[#tempPositionOfPrePostfix + 1] = #LGCODE_MTH_PRSR_CLOSE_BRACKET) OR
       (#tempPrePostfix[#tempPositionOfPrePostfix + 1] = #LGCODE_MTH_PRSR_LOGICAL_GREATER_EQUAL) OR
       (#tempPrePostfix[#tempPositionOfPrePostfix + 1] = #LGCODE_MTH_PRSR_LOGICAL_LESS_EQUAL) OR
       (#tempPrePostfix[#tempPositionOfPrePostfix + 1] = #LGCODE_MTH_PRSR_LOGICAL_NOT_EQUAL) OR
       (#tempPrePostfix[#tempPositionOfPrePostfix + 1] = #LGCODE_MTH_PRSR_PLUS) OR
       (#tempPrePostfix[#tempPositionOfPrePostfix + 1] = #LGCODE_MTH_PRSR_MINUS) OR
       (#tempPrePostfix[#tempPositionOfPrePostfix + 1] = #LGCODE_MTH_PRSR_TIMES) OR
       (#tempPrePostfix[#tempPositionOfPrePostfix + 1] = #LGCODE_MTH_PRSR_DIVIDE) OR
       (#tempPrePostfix[#tempPositionOfPrePostfix + 1] = #LGCODE_MTH_PRSR_TO_THE_POWER_OF) OR
       (#tempPositionOfPrePostfix = #tempMaxPositionOfPrePostfix))
     THEN
       IF (#tempDecimalPoint > 1) THEN
         #tempDecimalPoint := #tempDecimalPoint - 1;
       END_IF;
       #tempNumberOfBrackets := #tempNumberOfBrackets - 1;
     ELSE    //Falls keine der zulaessigen Kombinationen erfüllt ist
       #LKinLang_CalcMathAndBool.errorID := #LGCODE_MTH_PRSR_ERR_ID_INVALID_SYNTAX;
       #LKinLang_CalcMathAndBool.finalResult := 0;

       RETURN;
     END_IF;
     IF (#tempDecimalPoint > 2) OR (#tempNumberOfBrackets < 1) THEN    //Falls mehr als ein Komma pro Zahl
       #LKinLang_CalcMathAndBool.errorID := #LGCODE_MTH_PRSR_ERR_ID_INVALID_SYNTAX;
       #LKinLang_CalcMathAndBool.finalResult := 0;

       RETURN;
     END_IF;
     #tempPositionOfPrePostfix := #tempPositionOfPrePostfix + 1;
   END_WHILE;

   IF (#tempNumberOfBrackets <> 1) THEN    //Falls die Anzahl der Klammern nicht stimmt
     #LKinLang_CalcMathAndBool.errorID := #LGCODE_MTH_PRSR_ERR_ID_INVALID_SYNTAX;
     #LKinLang_CalcMathAndBool.finalResult := 0;

     RETURN;
   END_IF;
   #tempPositionOfPrePostfix := 1;

   //Beginn Umformung in Postfix-Notation
   WHILE #tempPositionOfPrePostfix <= #tempMaxPositionOfPrePostfix DO
     IF
       //Wenn Zahl und danach Dezimalpunkt, Dezimalzahl erzeugen
       (#tempPrePostfix[#tempPositionOfPrePostfix] <= #LGCODE_MTH_PRSR_NUMBER_9) AND
       (#tempPrePostfix[#tempPositionOfPrePostfix] >= #LGCODE_MTH_PRSR_NUMBER_0) AND
       (#tempPrePostfix[#tempPositionOfPrePostfix + 1] = #LGCODE_MTH_PRSR_DECIMAL_POINT)
     THEN
       #tempPostfixNotation[#tempPositionOfPostfix] := (#tempPrePostfix[#tempPositionOfPrePostfix] - #LGCODE_MTH_PRSR_NUMBER_0);

